screen "RIO 1 Analogue Settings" 1280x800, template "Template"
   on GenerateScreen: "TitleUpdater"()
   Button "HmiScreenItemData_1" at 1,1 size 150x40; TextOn 'Back'; TextOff 'Commissioning'
      on Release: ActivateScreen("Commissioning Main Page", 0)
   TextField "Text field_82" at 60,138 size 215x20; Text 'FPT USD Flow FIT-418-FPT'
   TextField "Text field_90" at 286,114 size 62x18; Text 'Reading'
   IOField "I/O field_2" at 281,138 size 75x20; FormatPattern 999; Unit  Nm³/hr
      ProcessValue <- "20_TANKS_IP_DATA_RIO_01_FIRST_TANK_USD_FLOW"
   TextField "Text field_1" at 359,114 size 68x18; Text 'Low Low'
   IOField "I/O field_1" at 361,138 size 60x20; Authorization "User administration"; FormatPattern 999
      ProcessValue <- "2084_Setpoints_FIT418_LoLo"
   TextField "Text field_2" at 442,114 size 34x18; Text 'Low'
   IOField "I/O field_3" at 429,138 size 60x20; Authorization "User administration"; FormatPattern 999
      ProcessValue <- "2084_Setpoints_FIT418_Lo"
   TextField "Text field_3" at 509,114 size 37x18; Text 'High'
   IOField "I/O field_4" at 497,138 size 60x20; Authorization "User administration"; FormatPattern 999
      ProcessValue <- "2084_Setpoints_FIT418_Hi"
   TextField "Text field_4" at 561,114 size 74x18; Text 'High High'
   IOField "I/O field_5" at 565,138 size 60x20; Authorization "User administration"; FormatPattern 999
      ProcessValue <- "2084_Setpoints_FIT418_HiHi"
   TextField "Text field_5" at 434,92 size 74x18; Text 'Setpoints'
   TextField "Text field_6" at 7,138 size 53x20; Text 'IW100'
   TextField "Text field_7" at 60,175 size 215x20; Text 'FPT MBG Flow FIT-420-FPT'
   IOField "I/O field_6" at 281,175 size 75x20; FormatPattern 999; Unit  Nm³/hr
      ProcessValue <- "20_TANKS_IP_DATA_RIO_01_FIRST_TANK_MBG_FLOW"
   IOField "I/O field_7" at 361,175 size 60x20; FormatPattern 999
      ProcessValue <- "2084_Setpoints_FIT420_LoLo"
   IOField "I/O field_8" at 429,175 size 60x20; FormatPattern 999
      ProcessValue <- "2084_Setpoints_FIT420_Lo"
   IOField "I/O field_9" at 497,175 size 60x20; Authorization "User administration"; FormatPattern 999
      ProcessValue <- "2084_Setpoints_FIT420_Hi"
   IOField "I/O field_10" at 565,175 size 60x20; Authorization "User administration"; FormatPattern 999
      ProcessValue <- "2084_Setpoints_FIT420_HiHi"
   TextField "Text field_8" at 7,175 size 53x20; Text 'IW102'
   TextField "Text field_9" at 60,212 size 215x20; Text 'Tank 1P USD Flow FIT-418-1P'
   IOField "I/O field_11" at 281,212 size 75x20; FormatPattern 999; Unit  Nm³/hr
      ProcessValue <- "20_TANKS_IP_DATA_RIO_01_SECOND_TANK_USD_FLOW"
   IOField "I/O field_12" at 361,212 size 60x20; FormatPattern 999
      ProcessValue <- "2084_Setpoints_FIT418_LoLo"
   IOField "I/O field_13" at 429,212 size 60x20; FormatPattern 999
      ProcessValue <- "2084_Setpoints_FIT418_Lo"
   IOField "I/O field_14" at 497,212 size 60x20; Authorization "User administration"; FormatPattern 999
      ProcessValue <- "2084_Setpoints_FIT418_Hi"
   IOField "I/O field_15" at 565,212 size 60x20; Authorization "User administration"; FormatPattern 999
      ProcessValue <- "2084_Setpoints_FIT418_HiHi"
   TextField "Text field_10" at 7,212 size 53x20; Text 'IW104'
   TextField "Text field_11" at 60,249 size 215x20; Text 'Tank 1P MBG Flow FIT-420-1P'
   IOField "I/O field_16" at 281,249 size 75x20; FormatPattern 999; Unit  Nm³/hr
      ProcessValue <- "20_TANKS_IP_DATA_RIO_01_SECOND_TANK_MBG_FLOW"
   IOField "I/O field_17" at 361,249 size 60x20; FormatPattern 999
      ProcessValue <- "2084_Setpoints_FIT420_LoLo"
   IOField "I/O field_18" at 429,249 size 60x20; FormatPattern 999
      ProcessValue <- "2084_Setpoints_FIT420_Lo"
   IOField "I/O field_19" at 497,249 size 60x20; FormatPattern 999
      ProcessValue <- "2084_Setpoints_FIT420_Hi"
   IOField "I/O field_20" at 565,249 size 60x20; FormatPattern 999
      ProcessValue <- "2084_Setpoints_FIT420_HiHi"
   TextField "Text field_12" at 7,249 size 53x20; Text 'IW106'
   TextField "Text field_13" at 60,286 size 215x20; Text 'Tank 1S USD Flow FIT-417-1S'
   IOField "I/O field_21" at 281,286 size 75x20; FormatPattern 999; Unit  Nm³/hr
      ProcessValue <- "20_TANKS_IP_DATA_RIO_01_THIRD_TANK_USD_FLOW"
   TextField "Text field_14" at 7,286 size 53x20; Text 'IW108'
   TextField "Text field_15" at 60,324 size 215x20; Text 'Tank 1S MBG Flow FIT-419-1S'
   IOField "I/O field_26" at 281,324 size 75x20; FormatPattern 999; Unit  Nm³/hr
      ProcessValue <- "20_TANKS_IP_DATA_RIO_01_THIRD_TANK_MBG_FLOW"
   TextField "Text field_16" at 7,324 size 53x20; Text 'IW110'
   TextField "Text field_17" at 60,361 size 215x20; Text 'FPT Confined Space Oxygen Level'
   IOField "I/O field_31" at 281,361 size 75x20; FormatPattern 99.9; Unit  %
      ProcessValue <- "20_TANKS_IP_DATA_RIO_01_FIRST_TANK_O2_MONITOR"
   IOField "I/O field_32" at 361,361 size 60x20; FormatPattern 99.9
      ProcessValue <- "2084_Setpoints_Conf O2 Level Lo Lo"
   IOField "I/O field_33" at 429,361 size 60x20; FormatPattern 99.9
      ProcessValue <- "2084_Setpoints_Conf O2 Level Lo"
   IOField "I/O field_34" at 497,361 size 60x20; FormatPattern 9.9
   IOField "I/O field_35" at 565,361 size 60x20; FormatPattern 9.9
   TextField "Text field_18" at 7,361 size 53x20; Text 'IW112'
   TextField "Text field_21" at 60,398 size 215x20; Text 'RIO 1 Deck Main Pressure PT-415'
   IOField "I/O field_41" at 281,398 size 75x20; FormatPattern 99.999; Unit  Bar
      ProcessValue <- "20_TANKS_IP_DATA_RIO_01_FIRST_TANK_DECK_IG_PRESS"
   IOField "I/O field_42" at 361,398 size 60x20; FormatPattern 99.99
      ProcessValue <- "2084_Setpoints_PIT415_LoLo"
   IOField "I/O field_43" at 429,398 size 60x20; FormatPattern 99.99
      ProcessValue <- "2084_Setpoints_PIT415_Lo"
   IOField "I/O field_44" at 497,398 size 60x20; FormatPattern 99.99
      ProcessValue <- "2084_Setpoints_PIT415_Hi"
   IOField "I/O field_45" at 565,398 size 60x20; FormatPattern 99.99
      ProcessValue <- "2084_Setpoints_PIT415_HiHi"
   TextField "Text field_22" at 7,398 size 53x20; Text 'IW116'
   TextField "Text field_23" at 60,435 size 215x20; Text 'FPT BW Level LT-422-FPT'
   IOField "I/O field_46" at 281,435 size 75x20; FormatPattern 999.9; Unit  %
      ProcessValue <- "20_TANKS_IP_DATA_RIO_01_FIRST_TANK_BWT_LEVEL"
   TextField "Text field_24" at 7,435 size 53x20; Text 'IW118'
   TextField "Text field_25" at 702,289 size 215x20; Text 'Tank 1P BW Temperature 426-1P'
   TextField "Text field_26" at 928,114 size 62x18; Text 'Reading'
   IOField "I/O field_51" at 922,289 size 75x20; FormatPattern s999.9; Unit  °C
      ProcessValue <- "20_TANKS_IP_DATA_RIO_01_SECOND_TANK_BWT_TEMP"
   TextField "Text field_27" at 1001,114 size 68x18; Text 'Low Low'
   TextField "Text field_28" at 1082,114 size 34x18; Text 'Low'
   TextField "Text field_29" at 1150,114 size 37x18; Text 'High'
   TextField "Text field_30" at 1203,114 size 74x18; Text 'High High'
   TextField "Text field_31" at 1076,92 size 74x18; Text 'Setpoints'
   TextField "Text field_32" at 649,289 size 53x20; Text 'IW150'
   TextField "Text field_33" at 702,326 size 215x20; Text 'Tank 1P BW DO TX-428-1P'
   IOField "I/O field_56" at 922,326 size 75x20; FormatPattern 99.9; Unit  mg/l
      ProcessValue <- "20_TANKS_IP_DATA_RIO_01_SECOND_TANK_BWT_DO"
   TextField "Text field_34" at 649,326 size 53x20; Text 'IW152'
   TextField "Text field_51" at 60,472 size 215x20; Text 'Tank 1P BW Level LT-422-1P'
   IOField "I/O field_101" at 281,472 size 75x20; FormatPattern 999.9; Unit  %
      ProcessValue <- "20_TANKS_IP_DATA_RIO_01_SECOND_TANK_BWT_LEVEL"
   TextField "Text field_56" at 7,472 size 53x20; Text 'IW120'
   TextField "Text field_57" at 60,509 size 215x20; Text 'Tank 1S BW Level LT-421-1S'
   IOField "I/O field_106" at 281,509 size 75x20; FormatPattern 999.9; Unit  %
      ProcessValue <- "20_TANKS_IP_DATA_RIO_01_THIRD_TANK_BWT_LEVEL"
   TextField "Text field_58" at 7,509 size 53x20; Text 'IW122'
   TextField "Text field_59" at 60,546 size 215x20; Text 'FPT BW ph TX-426-FPT'
   IOField "I/O field_111" at 281,546 size 75x20; FormatPattern 99.9
      ProcessValue <- "20_TANKS_IP_DATA_RIO_01_FIRST_TANK_BWT_PH"
   IOField "I/O field_112" at 361,546 size 60x20; FormatPattern 99.9
   IOField "I/O field_113" at 429,546 size 60x20; FormatPattern 99.9
      ProcessValue <- "2084_Setpoints_TX426 Port PH Lo"
   TextField "Text field_60" at 7,546 size 53x20; Text 'IW124'
   TextField "Text field_61" at 60,583 size 215x20; Text 'FPT BW Temperature 426-FPT'
   IOField "I/O field_116" at 281,583 size 75x20; FormatPattern 999.9; Unit  °C
      ProcessValue <- "20_TANKS_IP_DATA_RIO_01_FIRST_TANK_BWT_TEMP"
   IOField "I/O field_117" at 361,583 size 60x20; FormatPattern 99.9
   IOField "I/O field_118" at 429,583 size 60x20; FormatPattern 99.9
   TextField "Text field_62" at 7,583 size 53x20; Text 'IW126'
   TextField "Text field_63" at 60,620 size 215x20; Text 'FPT BW DO TX-428-FPT'
   IOField "I/O field_121" at 281,620 size 75x20; FormatPattern 99.9; Unit mg/l
      ProcessValue <- "20_TANKS_IP_DATA_RIO_01_FIRST_TANK_BWT_DO"
   TextField "Text field_64" at 7,620 size 53x20; Text 'IW128'
   TextField "Text field_65" at 702,138 size 215x20; Text 'Tank 1S BW ph TX-425-1S'
   IOField "I/O field_126" at 922,138 size 75x20; FormatPattern 99.9
      ProcessValue <- "20_TANKS_IP_DATA_RIO_01_THIRD_TANK_BWT_PH"
   TextField "Text field_66" at 649,138 size 53x20; Text 'IW140'
   TextField "Text field_67" at 702,175 size 215x20; Text 'Tank 1S BW Temperature 425-1S'
   IOField "I/O field_131" at 922,175 size 75x20; FormatPattern 999.9; Unit  °C
      ProcessValue <- "20_TANKS_IP_DATA_RIO_01_THIRD_TANK_BWT_TEMP"
   TextField "Text field_68" at 649,175 size 53x20; Text 'IW142'
   TextField "Text field_69" at 702,212 size 215x20; Text 'Tank 1S BW DO TX-427-1S'
   IOField "I/O field_136" at 922,212 size 75x20; FormatPattern 99.99; Unit  mg/l
      ProcessValue <- "20_TANKS_IP_DATA_RIO_01_THIRD_TANK_BWT_DO"
   TextField "Text field_70" at 649,212 size 53x20; Text 'IW144'
   TextField "Text field_73" at 702,251 size 215x20; Text 'Tank 1P BW ph TX-426-1P'
   IOField "I/O field_146" at 922,251 size 75x20; FormatPattern 99.9
      ProcessValue <- "20_TANKS_IP_DATA_RIO_01_SECOND_TANK_BWT_PH"
   TextField "Text field_74" at 649,251 size 53x20; Text 'IW148'
   TextField "Text field_41" at 133,114 size 85x18; Text 'Description'
   TextField "Text field_42" at 771,114 size 85x18; Text 'Description'
   TextField "Text field_43" at 17,114 size 21x18; Text 'AI'
   TextField "Text field_44" at 661,114 size 21x18; Text 'AI'
   TextField "Text field_47" at 59,657 size 215x20; Text 'RIO 1 Tanks Pressure PT-424'
   IOField "I/O field_81" at 280,657 size 75x20; FormatPattern s999.9; Unit  mBar
      ProcessValue <- "20_TANKS_IP_DATA_RIO_01_FIRST_TANK_TANKS_PRESS"
   TextField "Text field_48" at 6,657 size 53x20; Text 'IW130'
   IOField "I/O field_103" at 429,472 size 60x20; Authorization "User administration"; FormatPattern 999
      ProcessValue <- "2084_Setpoints_LT422_Lo"
   IOField "I/O field_104" at 497,472 size 60x20; Authorization "User administration"; FormatPattern 999
      ProcessValue <- "2084_Setpoints_LT422_Hi"
   IOField "I/O field_114" at 497,546 size 60x20; Authorization "User administration"; FormatPattern 99.9
      ProcessValue <- "2084_Setpoints_TX426 Port PH High"
   IOField "I/O field_115" at 565,546 size 60x20; Authorization "User administration"; FormatPattern 99.9
   IOField "I/O field_119" at 497,583 size 60x20; Authorization "User administration"; FormatPattern 99.9
   IOField "I/O field_120" at 565,583 size 60x20; Authorization "User administration"; FormatPattern 99.9
   IOField "I/O field_124" at 497,620 size 60x20; Authorization "User administration"; FormatPattern 99.9
      ProcessValue <- "2084_Setpoints_TX428 Port DO High"
   IOField "I/O field_125" at 565,620 size 60x20; Authorization "User administration"; FormatPattern 99.9
   IOField "I/O field_84" at 496,657 size 60x20; Authorization "User administration"; FormatPattern s999.9
      ProcessValue <- "2084_Setpoints_PIT424_Hi"
   IOField "I/O field_85" at 564,657 size 60x20; Authorization "User administration"; FormatPattern s999.9
      ProcessValue <- "2084_Setpoints_PIT424_HiHi"
   IOField "I/O field_122" at 361,620 size 60x20; Authorization "User administration"; FormatPattern 99.9
   IOField "I/O field_123" at 429,620 size 60x20; Authorization "User administration"; FormatPattern 99.9
      ProcessValue <- "2084_Setpoints_TX428 Port DO Lo"
   IOField "I/O field_82" at 360,657 size 60x20; Authorization "User administration"; FormatPattern s999.9
      ProcessValue <- "2084_Setpoints_PIT424_LoLo"
   IOField "I/O field_83" at 428,657 size 60x20; Authorization "User administration"; FormatPattern s999.9
      ProcessValue <- "2084_Setpoints_PIT424_Lo"
   IOField "I/O field_48" at 429,435 size 60x20; Authorization "User administration"; FormatPattern 999
      ProcessValue <- "2084_Setpoints_LT422_Lo"
   IOField "I/O field_49" at 497,435 size 60x20; Authorization "User administration"; FormatPattern 999
      ProcessValue <- "2084_Setpoints_LT422_Hi"
   IOField "I/O field_68" at 429,509 size 60x20; Authorization "User administration"; FormatPattern 999
      ProcessValue <- "2084_Setpoints_LT421_Lo"
   IOField "I/O field_69" at 497,509 size 60x20; Authorization "User administration"; FormatPattern 999
      ProcessValue <- "2084_Setpoints_LT421_Hi"
   IOField "I/O field_22" at 361,324 size 60x20; FormatPattern 999
      ProcessValue <- "2084_Setpoints_FIT419_LoLo"
   IOField "I/O field_23" at 429,324 size 60x20; FormatPattern 999
      ProcessValue <- "2084_Setpoints_FIT419_Lo"
   IOField "I/O field_24" at 497,324 size 60x20; FormatPattern 999
      ProcessValue <- "2084_Setpoints_FIT419_Hi"
   IOField "I/O field_25" at 565,324 size 60x20; FormatPattern 999
      ProcessValue <- "2084_Setpoints_FIT419_HiHi"
   IOField "I/O field_27" at 361,285 size 60x20; FormatPattern 999
      ProcessValue <- "2084_Setpoints_FIT417_LoLo"
   IOField "I/O field_28" at 429,285 size 60x20; FormatPattern 999
      ProcessValue <- "2084_Setpoints_FIT417_Lo"
   IOField "I/O field_29" at 497,285 size 60x20; Authorization "User administration"; FormatPattern 999
      ProcessValue <- "2084_Setpoints_FIT417_Hi"
   IOField "I/O field_30" at 565,285 size 60x20; Authorization "User administration"; FormatPattern 999
      ProcessValue <- "2084_Setpoints_FIT417_HiHi"
   IOField "I/O field_72" at 1003,251 size 60x20; FormatPattern 99.9
   IOField "I/O field_73" at 1071,251 size 60x20; FormatPattern 99.9
      ProcessValue <- "2084_Setpoints_TX426 Port PH Lo"
   IOField "I/O field_74" at 1003,289 size 60x20; FormatPattern 99.9
   IOField "I/O field_75" at 1071,289 size 60x20; FormatPattern 99.9
   IOField "I/O field_76" at 1139,251 size 60x20; Authorization "User administration"; FormatPattern 99.9
      ProcessValue <- "2084_Setpoints_TX426 Port PH High"
   IOField "I/O field_77" at 1207,251 size 60x20; Authorization "User administration"; FormatPattern 99.9
   IOField "I/O field_78" at 1139,289 size 60x20; Authorization "User administration"; FormatPattern 99.9
   IOField "I/O field_79" at 1207,289 size 60x20; Authorization "User administration"; FormatPattern 99.9
   IOField "I/O field_80" at 1139,326 size 60x20; Authorization "User administration"; FormatPattern 99.99
      ProcessValue <- "2084_Setpoints_TX428 Port DO High"
   IOField "I/O field_86" at 1207,326 size 60x20; Authorization "User administration"; FormatPattern 99.9
   IOField "I/O field_87" at 1003,326 size 60x20; Authorization "User administration"; FormatPattern 99.9
   IOField "I/O field_88" at 1071,326 size 60x20; Authorization "User administration"; FormatPattern 99.99
      ProcessValue <- "2084_Setpoints_TX428 Port DO Lo"
   IOField "I/O field_52" at 1003,138 size 60x20; FormatPattern 99.9
   IOField "I/O field_53" at 1071,138 size 60x20; FormatPattern 99.9
      ProcessValue <- "2084_Setpoints_TX425 Star PH Lo"
   IOField "I/O field_54" at 1003,175 size 60x20; FormatPattern 99.9
   IOField "I/O field_55" at 1071,175 size 60x20; FormatPattern 99.9
   IOField "I/O field_57" at 1139,138 size 60x20; Authorization "User administration"; FormatPattern 99.9
      ProcessValue <- "2084_Setpoints_TX425 Star PH High"
   IOField "I/O field_58" at 1207,138 size 60x20; Authorization "User administration"; FormatPattern 99.9
   IOField "I/O field_59" at 1139,175 size 60x20; Authorization "User administration"; FormatPattern 99.9
   IOField "I/O field_60" at 1207,175 size 60x20; Authorization "User administration"; FormatPattern 99.9
   IOField "I/O field_89" at 1139,212 size 60x20; Authorization "User administration"; FormatPattern 99.99
      ProcessValue <- "2084_Setpoints_TX427 Star DO High"
   IOField "I/O field_90" at 1207,212 size 60x20; Authorization "User administration"; FormatPattern 99.9
   IOField "I/O field_91" at 1003,212 size 60x20; Authorization "User administration"; FormatPattern 99.9
   IOField "I/O field_92" at 1071,212 size 60x20; Authorization "User administration"; FormatPattern 99.99
      ProcessValue <- "2084_Setpoints_TX427 Star DO Lo"
   IOField "I/O field_47" at 361,435 size 60x20; FormatPattern 9.9
   IOField "I/O field_66" at 361,472 size 60x20; FormatPattern 9.9
   IOField "I/O field_67" at 361,509 size 60x20; FormatPattern 9.9
   IOField "I/O field_50" at 565,435 size 60x20; FormatPattern 9.9
   IOField "I/O field_70" at 565,472 size 60x20; FormatPattern 9.9
   IOField "I/O field_71" at 565,509 size 60x20; FormatPattern 9.9
   Button "HmiScreenItemData_8" at 469,45 size 355x40; TextOn 'Back'; TextOff 'Text'
   TextField "Screen title" at 455,41 size 373x50; Text 'Screen title'

screen "RIO 2 Analogue Settings" 1280x800, template "Template"
   on GenerateScreen: "TitleUpdater"()
   Button "HmiScreenItemData_1" at 1,1 size 150x40; TextOn 'Back'; TextOff 'Commissioning'
      on Release: ActivateScreen("Commissioning Main Page", 0)
   TextField "Text field_82" at 60,138 size 215x20; Text 'Tank 2P USD Flow FIT-418-2P'
   TextField "Text field_90" at 286,114 size 62x18; Text 'Reading'
   IOField "I/O field_2" at 281,138 size 75x20; FormatPattern 999; Unit  Nm³/hr
      ProcessValue <- "20_TANKS_IP_DATA_RIO_02_FIRST_TANK_USD_FLOW"
   TextField "Text field_1" at 359,114 size 68x18; Text 'Low Low'
   TextField "Text field_2" at 442,114 size 34x18; Text 'Low'
   TextField "Text field_3" at 509,114 size 37x18; Text 'High'
   TextField "Text field_4" at 561,114 size 74x18; Text 'High High'
   TextField "Text field_5" at 434,92 size 74x18; Text 'Setpoints'
   TextField "Text field_6" at 7,138 size 53x20; Text 'IW160'
   TextField "Text field_7" at 60,175 size 215x20; Text 'Tank 2P MBG Flow FIT-420-2P'
   IOField "I/O field_6" at 281,175 size 75x20; FormatPattern 999; Unit  Nm³/hr
      ProcessValue <- "20_TANKS_IP_DATA_RIO_02_FIRST_TANK_MBG_FLOW"
   TextField "Text field_8" at 7,175 size 53x20; Text 'IW162'
   TextField "Text field_9" at 60,212 size 215x20; Text 'Tank 2S USD Flow FIT-417-2S'
   IOField "I/O field_11" at 281,212 size 75x20; FormatPattern 999; Unit  Nm³/hr
      ProcessValue <- "20_TANKS_IP_DATA_RIO_02_SECOND_TANK_USD_FLOW"
   TextField "Text field_10" at 7,212 size 53x20; Text 'IW164'
   TextField "Text field_11" at 60,249 size 215x20; Text 'Tank 2S MBG Flow FIT-419-2S'
   IOField "I/O field_16" at 281,249 size 75x20; FormatPattern 999; Unit  Nm³/hr
      ProcessValue <- "20_TANKS_IP_DATA_RIO_02_SECOND_TANK_MBG_FLOW"
   TextField "Text field_12" at 7,249 size 53x20; Text 'IW166'
   TextField "Text field_13" at 60,286 size 215x20; Text 'RIO 2 Deck Main Pressure PT-415'
   TextField "Text field_14" at 7,286 size 53x20; Text 'IW168'
   TextField "Text field_15" at 60,324 size 215x20; Text 'Tank 2P BW Level LT-422-2P'
   TextField "Text field_16" at 7,324 size 53x20; Text 'IW170'
   TextField "Text field_17" at 60,361 size 215x20; Text 'Tank 2S BW Level LT-421-2S'
   TextField "Text field_18" at 7,361 size 53x20; Text 'IW172'
   TextField "Text field_25" at 702,324 size 215x20; Text 'Tank 2S BW Temperature 425-2S'
   TextField "Text field_26" at 928,114 size 62x18; Text 'Reading'
   IOField "I/O field_51" at 922,324 size 75x20; FormatPattern s999.9; Unit  °C
      ProcessValue <- "20_TANKS_IP_DATA_RIO_02_SECOND_TANK_BWT_TEMP"
   TextField "Text field_27" at 1001,114 size 68x18; Text 'Low Low'
   TextField "Text field_28" at 1082,114 size 34x18; Text 'Low'
   TextField "Text field_29" at 1150,114 size 37x18; Text 'High'
   TextField "Text field_30" at 1203,114 size 74x18; Text 'High High'
   TextField "Text field_31" at 1076,92 size 74x18; Text 'Setpoints'
   TextField "Text field_32" at 649,324 size 53x20; Text 'IW186'
   TextField "Text field_33" at 702,361 size 215x20; Text 'Tank 2S BW DO TX-427-2S'
   IOField "I/O field_56" at 922,361 size 75x20; FormatPattern s99.99; Unit  mg/l
      ProcessValue <- "20_TANKS_IP_DATA_RIO_02_SECOND_TANK_BWT_DO"
   TextField "Text field_34" at 649,361 size 53x20; Text 'IW188'
   TextField "Text field_35" at 702,398 size 215x20; Text 'Confined Space O2 Level Port'
   TextField "Text field_36" at 649,398 size 53x20; Text 'IW190'
   TextField "Text field_65" at 702,138 size 215x20; Text 'Tank 2P BW ph TX-426-2P'
   IOField "I/O field_126" at 922,138 size 75x20; FormatPattern 99.9
      ProcessValue <- "20_TANKS_IP_DATA_RIO_02_FIRST_TANK_BWT_PH"
   TextField "Text field_66" at 649,138 size 53x20; Text 'IW176'
   TextField "Text field_67" at 702,175 size 215x20; Text 'Tank 2P BW Temperature 426-2P'
   IOField "I/O field_131" at 922,175 size 75x20; FormatPattern s999.9; Unit  °C
      ProcessValue <- "20_TANKS_IP_DATA_RIO_02_FIRST_TANK_BWT_TEMP"
   TextField "Text field_68" at 649,175 size 53x20; Text 'IW178'
   TextField "Text field_69" at 702,212 size 215x20; Text 'Tank 2P BW DO TX-428-2P'
   IOField "I/O field_136" at 922,212 size 75x20; FormatPattern s99.99; Unit  mg/l
      ProcessValue <- "20_TANKS_IP_DATA_RIO_02_FIRST_TANK_BWT_DO"
   TextField "Text field_70" at 649,212 size 53x20; Text 'IW180'
   TextField "Text field_71" at 702,249 size 215x20; Text 'RIO 2 Tanks Pressure PT-424'
   TextField "Text field_72" at 649,249 size 53x20; Text 'IW182'
   TextField "Text field_73" at 702,286 size 215x20; Text 'Tank 2S BW ph TX-425-2S'
   IOField "I/O field_146" at 922,286 size 75x20; FormatPattern 99.9
      ProcessValue <- "20_TANKS_IP_DATA_RIO_02_SECOND_TANK_BWT_PH"
   TextField "Text field_74" at 649,286 size 53x20; Text 'IW184'
   TextField "Text field_41" at 133,114 size 85x18; Text 'Description'
   TextField "Text field_42" at 771,114 size 85x18; Text 'Description'
   TextField "Text field_43" at 17,114 size 21x18; Text 'AI'
   TextField "Text field_44" at 661,114 size 21x18; Text 'AI'
   IOField "I/O field_21" at 281,285 size 75x20; FormatPattern 99.999; Unit  Bar
      ProcessValue <- "20_TANKS_IP_DATA_RIO_02_FIRST_TANK_DECK_IG_PRESS"
   IOField "I/O field_26" at 281,322 size 75x20; FormatPattern 999.9; Unit  %
      ProcessValue <- "20_TANKS_IP_DATA_RIO_02_FIRST_TANK_BWT_LEVEL"
   IOField "I/O field_27" at 281,359 size 75x20; FormatPattern 999.9; Unit  %
      ProcessValue <- "20_TANKS_IP_DATA_RIO_02_SECOND_TANK_BWT_LEVEL"
   IOField "I/O field_93" at 922,249 size 75x20; FormatPattern s999.9; Unit  mBar
      ProcessValue <- "20_TANKS_IP_DATA_RIO_02_FIRST_TANK_TANKS_PRESS"
   IOField "I/O field_41" at 922,398 size 75x20; FormatPattern 99.9; Unit  %
      ProcessValue <- "20_TANKS_IP_DATA_RIO_02_FIRST_TANK_O2_MONITOR"
   TextField "Text field_21" at 703,437 size 215x20; Text 'Confined Space O2 Level Starboard'
   TextField "Text field_22" at 650,437 size 53x20; Text 'IW190'
   IOField "I/O field_44" at 923,437 size 75x20; FormatPattern 99.9; Unit  %
      ProcessValue <- "20_TANKS_IP_DATA_RIO_02_SECOND_TANK_O2_MONITOR"
   IOField "I/O field_1" at 361,138 size 60x20; Authorization "User administration"; FormatPattern 999
      ProcessValue <- "2084_Setpoints_FIT418_LoLo"
   IOField "I/O field_3" at 429,138 size 60x20; Authorization "User administration"; FormatPattern 999
      ProcessValue <- "2084_Setpoints_FIT418_Lo"
   IOField "I/O field_4" at 497,138 size 60x20; Authorization "User administration"; FormatPattern 999
      ProcessValue <- "2084_Setpoints_FIT418_Hi"
   IOField "I/O field_5" at 565,138 size 60x20; Authorization "User administration"; FormatPattern 999
      ProcessValue <- "2084_Setpoints_FIT418_HiHi"
   IOField "I/O field_7" at 361,175 size 60x20; FormatPattern 999
      ProcessValue <- "2084_Setpoints_FIT420_LoLo"
   IOField "I/O field_8" at 429,175 size 60x20; FormatPattern 999
      ProcessValue <- "2084_Setpoints_FIT420_Lo"
   IOField "I/O field_9" at 497,175 size 60x20; Authorization "User administration"; FormatPattern 999
      ProcessValue <- "2084_Setpoints_FIT420_Hi"
   IOField "I/O field_10" at 565,175 size 60x20; Authorization "User administration"; FormatPattern 999
      ProcessValue <- "2084_Setpoints_FIT420_HiHi"
   IOField "I/O field_12" at 361,212 size 60x20; FormatPattern 999
      ProcessValue <- "2084_Setpoints_FIT417_LoLo"
   IOField "I/O field_13" at 429,212 size 60x20; FormatPattern 999
      ProcessValue <- "2084_Setpoints_FIT417_Lo"
   IOField "I/O field_14" at 497,212 size 60x20; Authorization "User administration"; FormatPattern 999
      ProcessValue <- "2084_Setpoints_FIT417_Hi"
   IOField "I/O field_15" at 565,212 size 60x20; Authorization "User administration"; FormatPattern 999
      ProcessValue <- "2084_Setpoints_FIT417_HiHi"
   IOField "I/O field_17" at 361,249 size 60x20; FormatPattern 999
      ProcessValue <- "2084_Setpoints_FIT419_LoLo"
   IOField "I/O field_18" at 429,249 size 60x20; FormatPattern 999
      ProcessValue <- "2084_Setpoints_FIT419_Lo"
   IOField "I/O field_19" at 497,249 size 60x20; FormatPattern 999
      ProcessValue <- "2084_Setpoints_FIT419_Hi"
   IOField "I/O field_20" at 565,249 size 60x20; FormatPattern 999
      ProcessValue <- "2084_Setpoints_FIT419_HiHi"
   IOField "I/O field_22" at 361,285 size 60x20; FormatPattern 99.999
      ProcessValue <- "2084_Setpoints_PIT415_LoLo"
   IOField "I/O field_23" at 429,285 size 60x20; FormatPattern 99.999
      ProcessValue <- "2084_Setpoints_PIT415_Lo"
   IOField "I/O field_24" at 497,285 size 60x20; FormatPattern 99.999
      ProcessValue <- "2084_Setpoints_PIT415_Hi"
   IOField "I/O field_25" at 565,285 size 60x20; FormatPattern 99.999
      ProcessValue <- "2084_Setpoints_PIT415_HiHi"
   IOField "I/O field_28" at 429,359 size 60x20; Authorization "User administration"; FormatPattern 999
      ProcessValue <- "2084_Setpoints_LT421_Lo"
   IOField "I/O field_29" at 497,359 size 60x20; Authorization "User administration"; FormatPattern 999
      ProcessValue <- "2084_Setpoints_LT421_Hi"
   IOField "I/O field_30" at 429,322 size 60x20; Authorization "User administration"; FormatPattern 999
      ProcessValue <- "2084_Setpoints_LT422_Lo"
   IOField "I/O field_31" at 497,322 size 60x20; Authorization "User administration"; FormatPattern 999
      ProcessValue <- "2084_Setpoints_LT422_Hi"
   IOField "I/O field_32" at 361,322 size 60x20; FormatPattern 9.9
   IOField "I/O field_33" at 361,359 size 60x20; FormatPattern 9.9
   IOField "I/O field_34" at 565,322 size 60x20; FormatPattern 9.9
   IOField "I/O field_35" at 565,359 size 60x20; FormatPattern 9.9
   IOField "I/O field_62" at 1004,397 size 60x20; FormatPattern 99.9
      ProcessValue <- "2084_Setpoints_Conf O2 Level Lo Lo"
   IOField "I/O field_63" at 1072,397 size 60x20; FormatPattern 99.9
      ProcessValue <- "2084_Setpoints_Conf O2 Level Lo"
   IOField "I/O field_64" at 1139,397 size 60x20; Authorization "User administration"; FormatPattern 99.9
   IOField "I/O field_65" at 1207,397 size 60x20; Authorization "User administration"; FormatPattern 99.9
   IOField "I/O field_72" at 1004,286 size 60x20; FormatPattern 99.9
   IOField "I/O field_74" at 1004,323 size 60x20; FormatPattern 99.9
   IOField "I/O field_75" at 1072,323 size 60x20; FormatPattern 99.9
   IOField "I/O field_77" at 1207,286 size 60x20; Authorization "User administration"; FormatPattern 99.9
   IOField "I/O field_78" at 1139,323 size 60x20; Authorization "User administration"; FormatPattern 99.9
   IOField "I/O field_79" at 1207,323 size 60x20; Authorization "User administration"; FormatPattern 99.9
   IOField "I/O field_80" at 1139,360 size 60x20; Authorization "User administration"; FormatPattern 99.9
      ProcessValue <- "2084_Setpoints_TX427 Star DO High"
   IOField "I/O field_86" at 1207,360 size 60x20; Authorization "User administration"; FormatPattern 99.9
   IOField "I/O field_87" at 1004,360 size 60x20; Authorization "User administration"; FormatPattern 99.9
   IOField "I/O field_88" at 1072,360 size 60x20; Authorization "User administration"; FormatPattern 99.9
      ProcessValue <- "2084_Setpoints_TX427 Star DO Lo"
   IOField "I/O field_52" at 1003,138 size 60x20; FormatPattern 99.9
   IOField "I/O field_53" at 1071,138 size 60x20; FormatPattern 99.9
      ProcessValue <- "2084_Setpoints_TX426 Port PH Lo"
   IOField "I/O field_54" at 1003,175 size 60x20; FormatPattern 99.9
   IOField "I/O field_55" at 1071,175 size 60x20; FormatPattern 99.9
   IOField "I/O field_57" at 1139,138 size 60x20; Authorization "User administration"; FormatPattern 99.9
      ProcessValue <- "2084_Setpoints_TX426 Port PH High"
   IOField "I/O field_58" at 1207,138 size 60x20; Authorization "User administration"; FormatPattern 99.9
   IOField "I/O field_59" at 1139,175 size 60x20; Authorization "User administration"; FormatPattern 99.9
   IOField "I/O field_60" at 1207,175 size 60x20; Authorization "User administration"; FormatPattern 99.9
   IOField "I/O field_89" at 1139,212 size 60x20; Authorization "User administration"; FormatPattern 99.9
      ProcessValue <- "2084_Setpoints_TX428 Port DO High"
   IOField "I/O field_90" at 1207,212 size 60x20; Authorization "User administration"; FormatPattern 99.9
   IOField "I/O field_91" at 1003,212 size 60x20; Authorization "User administration"; FormatPattern 99.9
   IOField "I/O field_92" at 1071,212 size 60x20; Authorization "User administration"; FormatPattern 99.9
      ProcessValue <- "2084_Setpoints_TX428 Port DO Lo"
   IOField "I/O field_94" at 1139,249 size 60x20; Authorization "User administration"; FormatPattern 999.9
      ProcessValue <- "2084_Setpoints_PIT424_Hi"
   IOField "I/O field_95" at 1207,249 size 60x20; Authorization "User administration"; FormatPattern 999.9
      ProcessValue <- "2084_Setpoints_PIT424_HiHi"
   IOField "I/O field_96" at 1004,249 size 60x20; Authorization "User administration"; FormatPattern 999.9
      ProcessValue <- "2084_Setpoints_PIT424_LoLo"
   IOField "I/O field_97" at 1072,249 size 60x20; Authorization "User administration"; FormatPattern 999.9
      ProcessValue <- "2084_Setpoints_PIT424_Lo"
   IOField "I/O field_42" at 1072,286 size 60x20; FormatPattern 99.9
      ProcessValue <- "2084_Setpoints_TX425 Star PH Lo"
   IOField "I/O field_43" at 1139,286 size 60x20; Authorization "User administration"; FormatPattern 99.9
      ProcessValue <- "2084_Setpoints_TX425 Star PH High"
   Button "HmiScreenItemData_8" at 469,45 size 355x40; TextOn 'Back'; TextOff 'Text'
   TextField "Screen title" at 455,41 size 373x50; Text 'Screen title'

screen "RIO 3 Analogue Settings" 1280x800, template "Template"
   on GenerateScreen: "TitleUpdater"()
   Button "HmiScreenItemData_1" at 1,1 size 150x40; TextOn 'Back'; TextOff 'Commissioning'
      on Release: ActivateScreen("Commissioning Main Page", 0)
   TextField "Text field_82" at 60,138 size 215x20; Text 'Tank 3P USD Flow FIT-418-3P'
   TextField "Text field_90" at 286,114 size 62x18; Text 'Reading'
   IOField "I/O field_2" at 281,138 size 75x20; FormatPattern 999; Unit  Nm³/hr
      ProcessValue <- "20_TANKS_IP_DATA_RIO_03_FIRST_TANK_USD_FLOW"
   TextField "Text field_1" at 359,114 size 68x18; Text 'Low Low'
   IOField "I/O field_1" at 361,138 size 60x20; Authorization "User administration"; FormatPattern 999
      ProcessValue <- "2084_Setpoints_FIT418_LoLo"
   TextField "Text field_2" at 442,114 size 34x18; Text 'Low'
   IOField "I/O field_3" at 429,138 size 60x20; Authorization "User administration"; FormatPattern 999
      ProcessValue <- "2084_Setpoints_FIT418_Lo"
   TextField "Text field_3" at 509,114 size 37x18; Text 'High'
   IOField "I/O field_4" at 497,138 size 60x20; Authorization "User administration"; FormatPattern 999
      ProcessValue <- "2084_Setpoints_FIT418_Hi"
   TextField "Text field_4" at 561,114 size 74x18; Text 'High High'
   IOField "I/O field_5" at 565,138 size 60x20; Authorization "User administration"; FormatPattern 999
      ProcessValue <- "2084_Setpoints_FIT418_HiHi"
   TextField "Text field_5" at 434,92 size 74x18; Text 'Setpoints'
   TextField "Text field_6" at 7,138 size 53x20; Text 'IW200'
   TextField "Text field_7" at 60,175 size 215x20; Text 'Tank 3P MBG Flow FIT-420-3P'
   IOField "I/O field_6" at 281,175 size 75x20; FormatPattern 999; Unit  Nm³/hr
      ProcessValue <- "20_TANKS_IP_DATA_RIO_03_FIRST_TANK_MBG_FLOW"
   IOField "I/O field_7" at 361,175 size 60x20; FormatPattern 999
      ProcessValue <- "2084_Setpoints_FIT420_LoLo"
   IOField "I/O field_8" at 429,175 size 60x20; FormatPattern 999
      ProcessValue <- "2084_Setpoints_FIT420_Lo"
   IOField "I/O field_9" at 497,175 size 60x20; Authorization "User administration"; FormatPattern 999
      ProcessValue <- "2084_Setpoints_FIT420_Hi"
   IOField "I/O field_10" at 565,175 size 60x20; Authorization "User administration"; FormatPattern 999
      ProcessValue <- "2084_Setpoints_FIT420_HiHi"
   TextField "Text field_8" at 7,175 size 53x20; Text 'IW202'
   TextField "Text field_9" at 60,212 size 215x20; Text 'Tank 3S USD Flow FIT-417-3S'
   IOField "I/O field_11" at 281,212 size 75x20; FormatPattern 999; Unit  Nm³/hr
      ProcessValue <- "20_TANKS_IP_DATA_RIO_03_SECOND_TANK_USD_FLOW"
   IOField "I/O field_12" at 361,212 size 60x20; FormatPattern 999
      ProcessValue <- "2084_Setpoints_FIT417_LoLo"
   IOField "I/O field_13" at 429,212 size 60x20; FormatPattern 999
      ProcessValue <- "2084_Setpoints_FIT417_Lo"
   IOField "I/O field_14" at 497,212 size 60x20; Authorization "User administration"; FormatPattern 999
      ProcessValue <- "2084_Setpoints_FIT417_Hi"
   IOField "I/O field_15" at 565,212 size 60x20; Authorization "User administration"; FormatPattern 999
      ProcessValue <- "2084_Setpoints_FIT417_HiHi"
   TextField "Text field_10" at 7,212 size 53x20; Text 'IW204'
   TextField "Text field_11" at 60,249 size 215x20; Text 'Tank 3S MBG Flow FIT-419-3S'
   IOField "I/O field_16" at 281,249 size 75x20; FormatPattern 999; Unit  Nm³/hr
      ProcessValue <- "20_TANKS_IP_DATA_RIO_03_SECOND_TANK_MBG_FLOW"
   IOField "I/O field_17" at 361,249 size 60x20; FormatPattern 999
      ProcessValue <- "2084_Setpoints_FIT419_LoLo"
   IOField "I/O field_18" at 429,249 size 60x20; FormatPattern 999
      ProcessValue <- "2084_Setpoints_FIT419_Lo"
   IOField "I/O field_19" at 497,249 size 60x20; FormatPattern 999
      ProcessValue <- "2084_Setpoints_FIT419_Hi"
   IOField "I/O field_20" at 565,249 size 60x20; FormatPattern 999
      ProcessValue <- "2084_Setpoints_FIT419_HiHi"
   TextField "Text field_12" at 7,249 size 53x20; Text 'IW206'
   TextField "Text field_13" at 60,286 size 215x20; Text 'RIO 3 Deck Main Pressure PT-415'
   TextField "Text field_14" at 7,286 size 53x20; Text 'IW208'
   TextField "Text field_15" at 60,324 size 215x20; Text 'Tank 3P BW Level LT-422-3P'
   TextField "Text field_16" at 7,324 size 53x20; Text 'IW210'
   TextField "Text field_17" at 60,361 size 215x20; Text 'Tank 3S BW Level LT-421-3S'
   TextField "Text field_18" at 7,361 size 53x20; Text 'IW212'
   TextField "Text field_25" at 702,323 size 215x20; Text 'Tank 3S BW Temperature 425-3S'
   TextField "Text field_26" at 928,114 size 62x18; Text 'Reading'
   IOField "I/O field_51" at 922,323 size 75x20; FormatPattern s999; Unit  °C
      ProcessValue <- "20_TANKS_IP_DATA_RIO_03_SECOND_TANK_BWT_TEMP"
   TextField "Text field_27" at 1001,114 size 68x18; Text 'Low Low'
   TextField "Text field_28" at 1082,114 size 34x18; Text 'Low'
   TextField "Text field_29" at 1150,114 size 37x18; Text 'High'
   TextField "Text field_30" at 1203,114 size 74x18; Text 'High High'
   TextField "Text field_31" at 1076,92 size 74x18; Text 'Setpoints'
   TextField "Text field_32" at 649,323 size 53x20; Text 'IW226'
   TextField "Text field_33" at 702,360 size 215x20; Text 'Tank 3S BW DO TX-427-3S'
   IOField "I/O field_56" at 922,360 size 75x20; FormatPattern 99.99; Unit  mg/l
      ProcessValue <- "20_TANKS_IP_DATA_RIO_03_SECOND_TANK_BWT_DO"
   TextField "Text field_34" at 649,360 size 53x20; Text 'IW228'
   TextField "Text field_35" at 702,397 size 215x20; Text 'Confined Space O2 Level Port'
   IOField "I/O field_61" at 922,397 size 75x20; FormatPattern 99.9; Unit  %
      ProcessValue <- "20_TANKS_IP_DATA_RIO_03_FIRST_TANK_O2_MONITOR"
   IOField "I/O field_62" at 1004,397 size 60x20; FormatPattern 99.9
      ProcessValue <- "2084_Setpoints_Conf O2 Level Lo Lo"
   IOField "I/O field_63" at 1072,397 size 60x20; FormatPattern 99.9
      ProcessValue <- "2084_Setpoints_Conf O2 Level Lo"
   TextField "Text field_36" at 649,397 size 53x20; Text 'IW230'
   TextField "Text field_65" at 702,138 size 215x20; Text 'Tank 3P BW ph TX-426-3P'
   IOField "I/O field_126" at 922,138 size 75x20; FormatPattern 99.9
      ProcessValue <- "20_TANKS_IP_DATA_RIO_03_FIRST_TANK_BWT_PH"
   TextField "Text field_66" at 649,138 size 53x20; Text 'IW216'
   TextField "Text field_67" at 702,175 size 215x20; Text 'Tank 3P BW Temperature 426-3P'
   IOField "I/O field_131" at 922,175 size 75x20; FormatPattern s999.9; Unit  °C
      ProcessValue <- "20_TANKS_IP_DATA_RIO_03_FIRST_TANK_BWT_TEMP"
   TextField "Text field_68" at 649,175 size 53x20; Text 'IW218'
   TextField "Text field_69" at 702,212 size 215x20; Text 'Tank 3P BW DO TX-428-3P'
   IOField "I/O field_136" at 922,212 size 75x20; FormatPattern 99.99; Unit  mg/l
      ProcessValue <- "20_TANKS_IP_DATA_RIO_03_FIRST_TANK_BWT_DO"
   TextField "Text field_70" at 649,212 size 53x20; Text 'IW220'
   TextField "Text field_71" at 702,249 size 215x20; Text 'RIO 3 Tanks Pressure PT-424'
   TextField "Text field_72" at 649,249 size 53x20; Text 'IW222'
   TextField "Text field_73" at 702,286 size 215x20; Text 'Tank 3S BW ph TX-425-3S'
   IOField "I/O field_146" at 922,286 size 75x20; FormatPattern 99.9
      ProcessValue <- "20_TANKS_IP_DATA_RIO_03_SECOND_TANK_BWT_PH"
   TextField "Text field_74" at 649,286 size 53x20; Text 'IW224'
   TextField "Text field_41" at 133,114 size 85x18; Text 'Description'
   TextField "Text field_42" at 771,114 size 85x18; Text 'Description'
   TextField "Text field_43" at 17,114 size 21x18; Text 'AI'
   TextField "Text field_44" at 661,114 size 21x18; Text 'AI'
   IOField "I/O field_64" at 1139,397 size 60x20; Authorization "User administration"; FormatPattern 99.9
   IOField "I/O field_65" at 1207,397 size 60x20; Authorization "User administration"; FormatPattern 99.9
   IOField "I/O field_72" at 1004,286 size 60x20; FormatPattern 99.9
   IOField "I/O field_74" at 1004,323 size 60x20; FormatPattern 99.9
   IOField "I/O field_75" at 1072,323 size 60x20; FormatPattern 99.9
   IOField "I/O field_77" at 1207,286 size 60x20; Authorization "User administration"; FormatPattern 99.9
   IOField "I/O field_78" at 1139,323 size 60x20; Authorization "User administration"; FormatPattern 99.9
   IOField "I/O field_79" at 1207,323 size 60x20; Authorization "User administration"; FormatPattern 99.9
   IOField "I/O field_80" at 1139,360 size 60x20; Authorization "User administration"; FormatPattern 99.9
      ProcessValue <- "2084_Setpoints_TX427 Star DO High"
   IOField "I/O field_86" at 1207,360 size 60x20; Authorization "User administration"; FormatPattern 99.9
   IOField "I/O field_87" at 1004,360 size 60x20; Authorization "User administration"; FormatPattern 99.9
   IOField "I/O field_88" at 1072,360 size 60x20; Authorization "User administration"; FormatPattern 99.9
      ProcessValue <- "2084_Setpoints_TX427 Star DO Lo"
   IOField "I/O field_52" at 1003,138 size 60x20; FormatPattern 99.9
   IOField "I/O field_53" at 1071,138 size 60x20; FormatPattern 99.9
      ProcessValue <- "2084_Setpoints_TX426 Port PH Lo"
   IOField "I/O field_54" at 1003,175 size 60x20; FormatPattern 99.9
   IOField "I/O field_55" at 1071,175 size 60x20; FormatPattern 99.9
   IOField "I/O field_57" at 1139,138 size 60x20; Authorization "User administration"; FormatPattern 99.9
      ProcessValue <- "2084_Setpoints_TX426 Port PH High"
   IOField "I/O field_58" at 1207,138 size 60x20; Authorization "User administration"; FormatPattern 99.9
   IOField "I/O field_59" at 1139,175 size 60x20; Authorization "User administration"; FormatPattern 99.9
   IOField "I/O field_60" at 1207,175 size 60x20; Authorization "User administration"; FormatPattern 99.9
   IOField "I/O field_89" at 1139,212 size 60x20; Authorization "User administration"; FormatPattern 99.9
      ProcessValue <- "2084_Setpoints_TX428 Port DO High"
   IOField "I/O field_90" at 1207,212 size 60x20; Authorization "User administration"; FormatPattern 99.9
   IOField "I/O field_91" at 1003,212 size 60x20; Authorization "User administration"; FormatPattern 99.9
   IOField "I/O field_92" at 1071,212 size 60x20; Authorization "User administration"; FormatPattern 99.9
      ProcessValue <- "2084_Setpoints_TX428 Port DO Lo"
   IOField "I/O field_21" at 281,285 size 75x20; FormatPattern 99.999; Unit  Bar
      ProcessValue <- "20_TANKS_IP_DATA_RIO_03_FIRST_TANK_DECK_IG_PRESS"
   IOField "I/O field_22" at 361,285 size 60x20; FormatPattern 99.999
      ProcessValue <- "2084_Setpoints_PIT415_LoLo"
   IOField "I/O field_23" at 429,285 size 60x20; FormatPattern 99.999
      ProcessValue <- "2084_Setpoints_PIT415_Lo"
   IOField "I/O field_24" at 497,285 size 60x20; FormatPattern 99.999
      ProcessValue <- "2084_Setpoints_PIT415_Hi"
   IOField "I/O field_25" at 565,285 size 60x20; FormatPattern 99.999
      ProcessValue <- "2084_Setpoints_PIT415_HiHi"
   IOField "I/O field_26" at 281,322 size 75x20; FormatPattern 999; Unit  %
      ProcessValue <- "20_TANKS_IP_DATA_RIO_03_FIRST_TANK_BWT_LEVEL"
   IOField "I/O field_27" at 281,359 size 75x20; FormatPattern 999.9; Unit  %
      ProcessValue <- "20_TANKS_IP_DATA_RIO_03_SECOND_TANK_BWT_LEVEL"
   IOField "I/O field_28" at 429,359 size 60x20; Authorization "User administration"; FormatPattern 999
      ProcessValue <- "2084_Setpoints_LT421_Lo"
   IOField "I/O field_29" at 497,359 size 60x20; Authorization "User administration"; FormatPattern 999
      ProcessValue <- "2084_Setpoints_LT421_Hi"
   IOField "I/O field_30" at 429,322 size 60x20; Authorization "User administration"; FormatPattern 999
      ProcessValue <- "2084_Setpoints_LT422_Lo"
   IOField "I/O field_31" at 497,322 size 60x20; Authorization "User administration"; FormatPattern 999
      ProcessValue <- "2084_Setpoints_LT422_Hi"
   IOField "I/O field_32" at 361,322 size 60x20; FormatPattern 9.9
   IOField "I/O field_33" at 361,359 size 60x20; FormatPattern 9.9
   IOField "I/O field_34" at 565,322 size 60x20; FormatPattern 9.9
   IOField "I/O field_35" at 565,359 size 60x20; FormatPattern 9.9
   IOField "I/O field_93" at 922,249 size 75x20; FormatPattern s99.9; Unit  mBar
      ProcessValue <- "20_TANKS_IP_DATA_RIO_03_FIRST_TANK_TANKS_PRESS"
   IOField "I/O field_94" at 1139,249 size 60x20; Authorization "User administration"; FormatPattern 999.9
      ProcessValue <- "2084_Setpoints_PIT424_Hi"
   IOField "I/O field_95" at 1207,249 size 60x20; Authorization "User administration"; FormatPattern 999.9
      ProcessValue <- "2084_Setpoints_PIT424_HiHi"
   IOField "I/O field_96" at 1004,249 size 60x20; Authorization "User administration"; FormatPattern 999.9
      ProcessValue <- "2084_Setpoints_PIT424_LoLo"
   IOField "I/O field_97" at 1072,249 size 60x20; Authorization "User administration"; FormatPattern 999.9
      ProcessValue <- "2084_Setpoints_PIT424_Lo"
   IOField "I/O field_41" at 1072,286 size 60x20; FormatPattern 99.9
      ProcessValue <- "2084_Setpoints_TX425 Star PH Lo"
   IOField "I/O field_42" at 1139,286 size 60x20; Authorization "User administration"; FormatPattern 99.9
      ProcessValue <- "2084_Setpoints_TX425 Star PH High"
   IOField "I/O field_43" at 922,435 size 75x20; FormatPattern 99.9; Unit  %
      ProcessValue <- "20_TANKS_IP_DATA_RIO_03_SECOND_TANK_O2_MONITOR"
   TextField "Text field_21" at 702,435 size 215x20; Text 'Confined Space O2 Level Starboard'
   TextField "Text field_22" at 649,435 size 53x20; Text 'IW230'
   Button "HmiScreenItemData_8" at 469,45 size 355x40; TextOn 'Back'; TextOff 'Text'
   TextField "Screen title" at 455,41 size 373x50; Text 'Screen title'